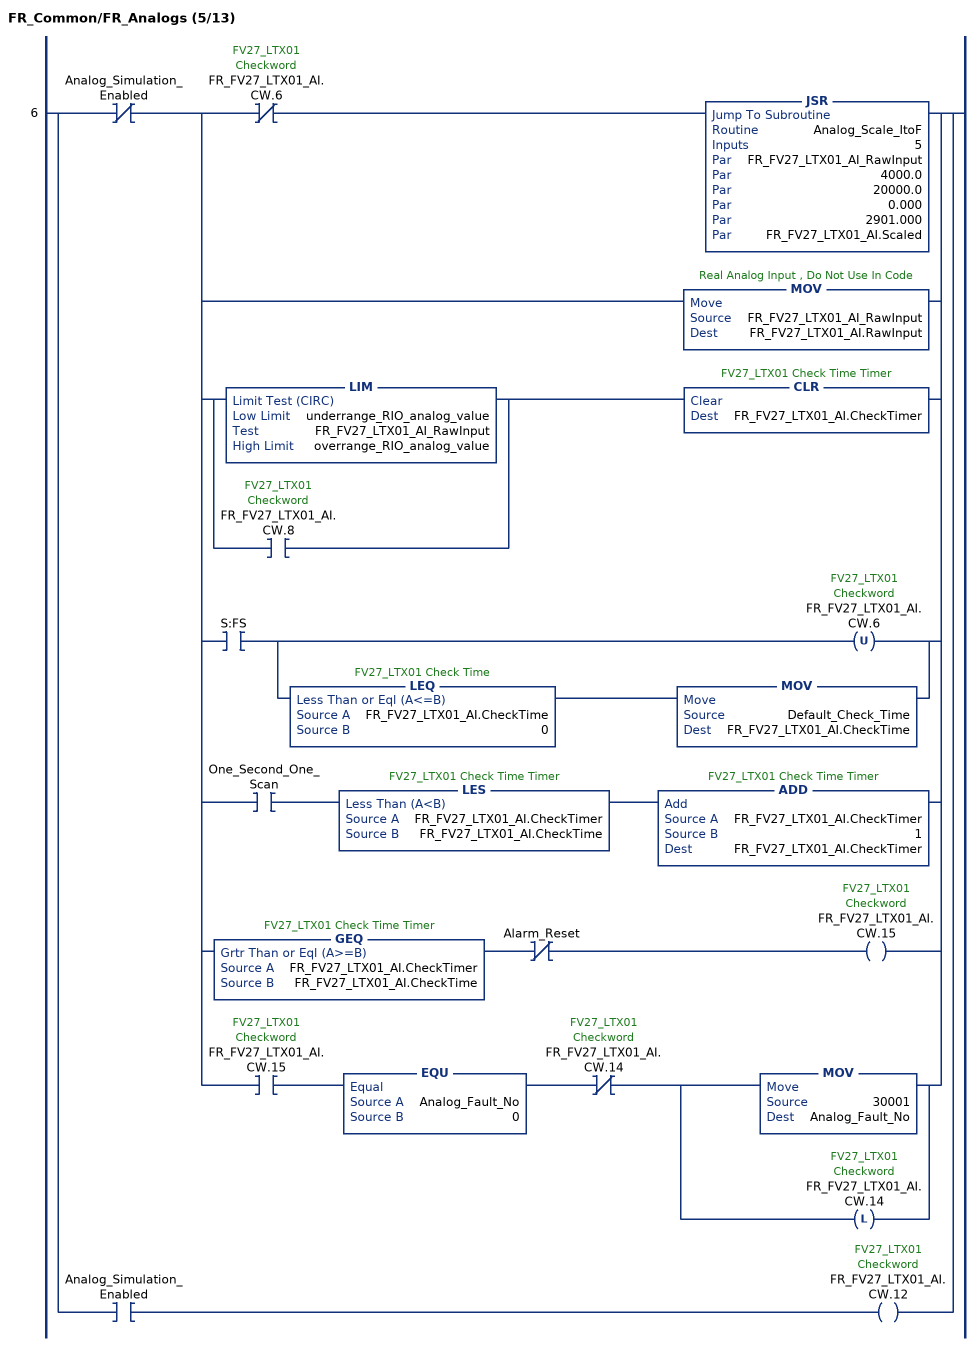
   6: [XIO(Analog_Simulation_Enabled) [XIO(FR_FV27_LTX01_AI.CW.6) JSR(Analog_Scale_ItoF,5,FR_FV27_LTX01_AI_RawInput,4000.0,20000.0,0.000,2901.000,FR_FV27_LTX01_AI.Scaled) ,MOV(FR_FV27_LTX01_AI_RawInput,FR_FV27_LTX01_AI.RawInput) ,[LIM(underrange_RIO_analog_value,FR_FV27_LTX01_AI_RawInput,overrange_RIO_analog_value) ,XIC(FR_FV27_LTX01_AI.CW.8) ] CLR(FR_FV27_LTX01_AI.CheckTimer) ,XIC(S:FS) [OTU(FR_FV27_LTX01_AI.CW.6) ,LEQ(FR_FV27_LTX01_AI.CheckTime,0) MOV(Default_Check_Time,FR_FV27_LTX01_AI.CheckTime) ] ,XIC(One_Second_One_Scan) LES(FR_FV27_LTX01_AI.CheckTimer,FR_FV27_LTX01_AI.CheckTime) ADD(FR_FV27_LTX01_AI.CheckTimer,1,FR_FV27_LTX01_AI.CheckTimer) ,GEQ(FR_FV27_LTX01_AI.CheckTimer,FR_FV27_LTX01_AI.CheckTime) XIO(Alarm_Reset) OTE(FR_FV27_LTX01_AI.CW.15) ,XIC(FR_FV27_LTX01_AI.CW.15) EQU(Analog_Fault_No,0) XIO(FR_FV27_LTX01_AI.CW.14) [MOV(30001,Analog_Fault_No) ,OTL(FR_FV27_LTX01_AI.CW.14) ] ] ,XIC(Analog_Simulation_Enabled) OTE(FR_FV27_LTX01_AI.CW.12) ];
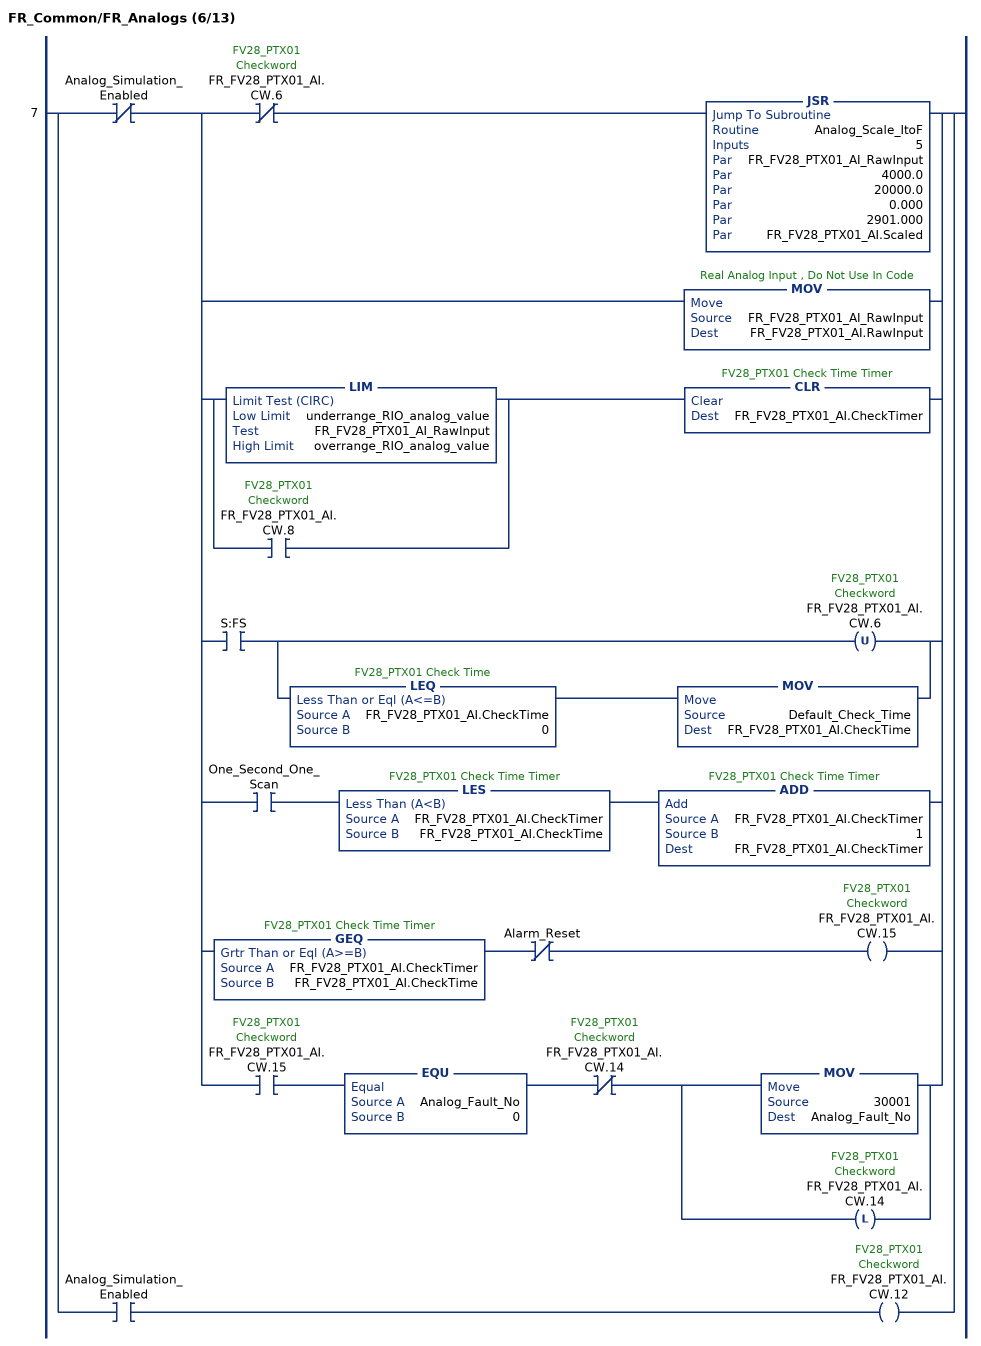
   7: [XIO(Analog_Simulation_Enabled) [XIO(FR_FV28_PTX01_AI.CW.6) JSR(Analog_Scale_ItoF,5,FR_FV28_PTX01_AI_RawInput,4000.0,20000.0,0.000,2901.000,FR_FV28_PTX01_AI.Scaled) ,MOV(FR_FV28_PTX01_AI_RawInput,FR_FV28_PTX01_AI.RawInput) ,[LIM(underrange_RIO_analog_value,FR_FV28_PTX01_AI_RawInput,overrange_RIO_analog_value) ,XIC(FR_FV28_PTX01_AI.CW.8) ] CLR(FR_FV28_PTX01_AI.CheckTimer) ,XIC(S:FS) [OTU(FR_FV28_PTX01_AI.CW.6) ,LEQ(FR_FV28_PTX01_AI.CheckTime,0) MOV(Default_Check_Time,FR_FV28_PTX01_AI.CheckTime) ] ,XIC(One_Second_One_Scan) LES(FR_FV28_PTX01_AI.CheckTimer,FR_FV28_PTX01_AI.CheckTime) ADD(FR_FV28_PTX01_AI.CheckTimer,1,FR_FV28_PTX01_AI.CheckTimer) ,GEQ(FR_FV28_PTX01_AI.CheckTimer,FR_FV28_PTX01_AI.CheckTime) XIO(Alarm_Reset) OTE(FR_FV28_PTX01_AI.CW.15) ,XIC(FR_FV28_PTX01_AI.CW.15) EQU(Analog_Fault_No,0) XIO(FR_FV28_PTX01_AI.CW.14) [MOV(30001,Analog_Fault_No) ,OTL(FR_FV28_PTX01_AI.CW.14) ] ] ,XIC(Analog_Simulation_Enabled) OTE(FR_FV28_PTX01_AI.CW.12) ];
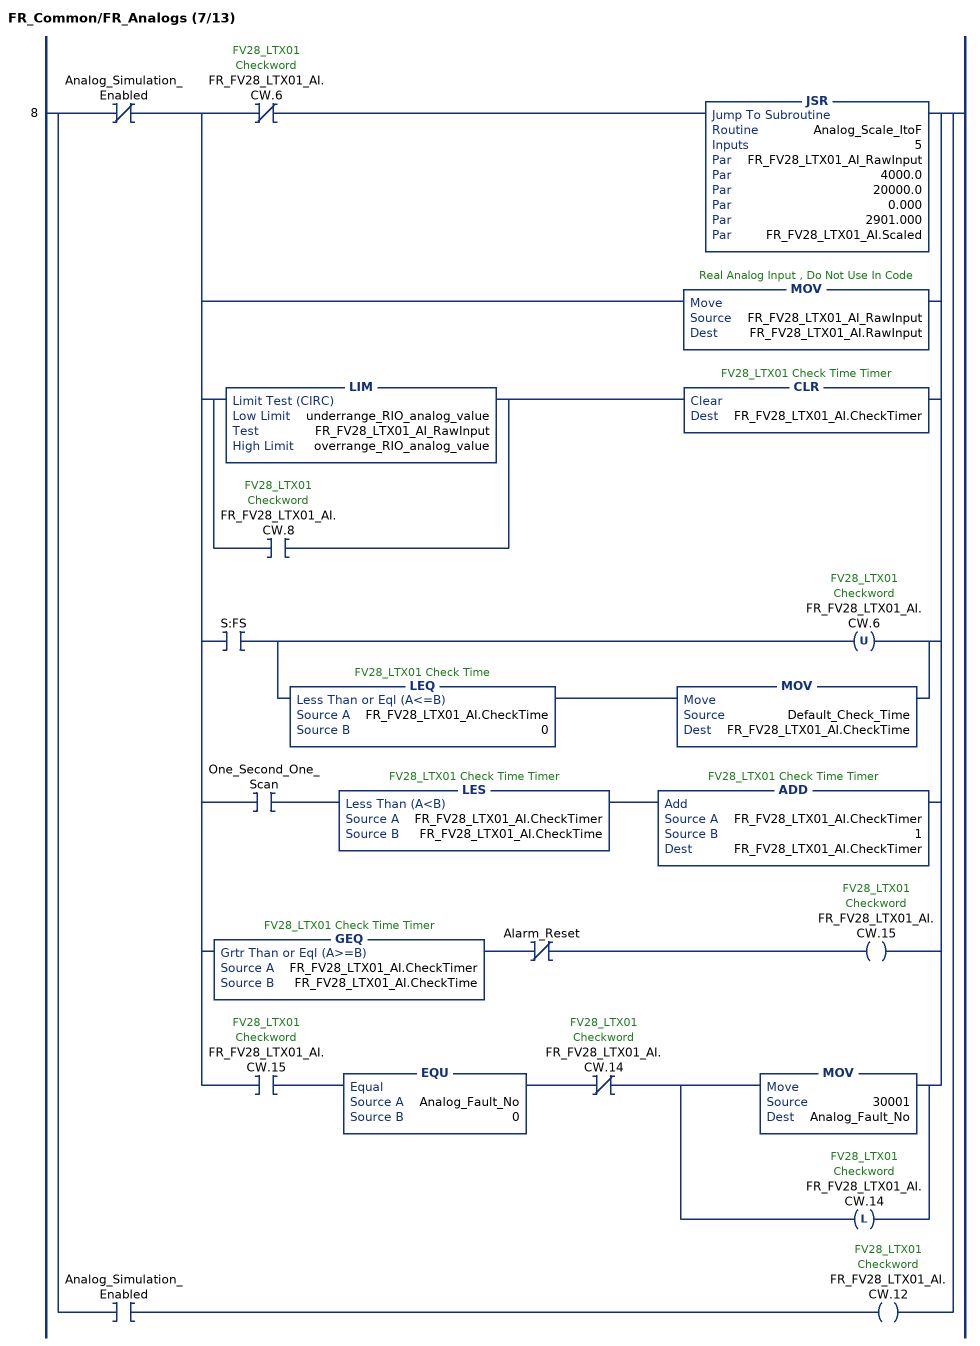
   8: [XIO(Analog_Simulation_Enabled) [XIO(FR_FV28_LTX01_AI.CW.6) JSR(Analog_Scale_ItoF,5,FR_FV28_LTX01_AI_RawInput,4000.0,20000.0,0.000,2901.000,FR_FV28_LTX01_AI.Scaled) ,MOV(FR_FV28_LTX01_AI_RawInput,FR_FV28_LTX01_AI.RawInput) ,[LIM(underrange_RIO_analog_value,FR_FV28_LTX01_AI_RawInput,overrange_RIO_analog_value) ,XIC(FR_FV28_LTX01_AI.CW.8) ] CLR(FR_FV28_LTX01_AI.CheckTimer) ,XIC(S:FS) [OTU(FR_FV28_LTX01_AI.CW.6) ,LEQ(FR_FV28_LTX01_AI.CheckTime,0) MOV(Default_Check_Time,FR_FV28_LTX01_AI.CheckTime) ] ,XIC(One_Second_One_Scan) LES(FR_FV28_LTX01_AI.CheckTimer,FR_FV28_LTX01_AI.CheckTime) ADD(FR_FV28_LTX01_AI.CheckTimer,1,FR_FV28_LTX01_AI.CheckTimer) ,GEQ(FR_FV28_LTX01_AI.CheckTimer,FR_FV28_LTX01_AI.CheckTime) XIO(Alarm_Reset) OTE(FR_FV28_LTX01_AI.CW.15) ,XIC(FR_FV28_LTX01_AI.CW.15) EQU(Analog_Fault_No,0) XIO(FR_FV28_LTX01_AI.CW.14) [MOV(30001,Analog_Fault_No) ,OTL(FR_FV28_LTX01_AI.CW.14) ] ] ,XIC(Analog_Simulation_Enabled) OTE(FR_FV28_LTX01_AI.CW.12) ];
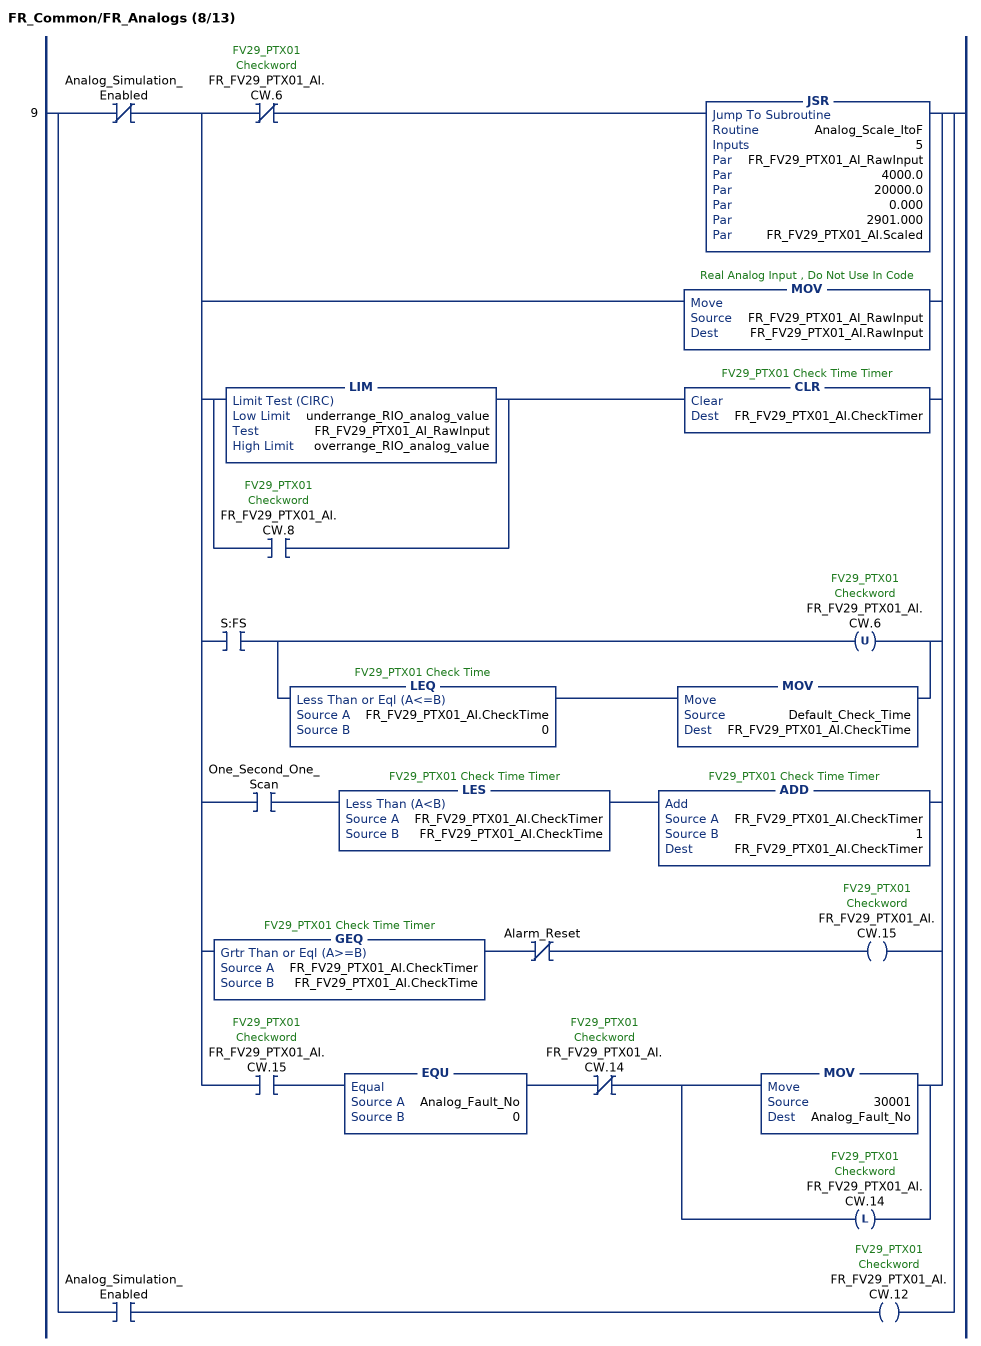
   9: [XIO(Analog_Simulation_Enabled) [XIO(FR_FV29_PTX01_AI.CW.6) JSR(Analog_Scale_ItoF,5,FR_FV29_PTX01_AI_RawInput,4000.0,20000.0,0.000,2901.000,FR_FV29_PTX01_AI.Scaled) ,MOV(FR_FV29_PTX01_AI_RawInput,FR_FV29_PTX01_AI.RawInput) ,[LIM(underrange_RIO_analog_value,FR_FV29_PTX01_AI_RawInput,overrange_RIO_analog_value) ,XIC(FR_FV29_PTX01_AI.CW.8) ] CLR(FR_FV29_PTX01_AI.CheckTimer) ,XIC(S:FS) [OTU(FR_FV29_PTX01_AI.CW.6) ,LEQ(FR_FV29_PTX01_AI.CheckTime,0) MOV(Default_Check_Time,FR_FV29_PTX01_AI.CheckTime) ] ,XIC(One_Second_One_Scan) LES(FR_FV29_PTX01_AI.CheckTimer,FR_FV29_PTX01_AI.CheckTime) ADD(FR_FV29_PTX01_AI.CheckTimer,1,FR_FV29_PTX01_AI.CheckTimer) ,GEQ(FR_FV29_PTX01_AI.CheckTimer,FR_FV29_PTX01_AI.CheckTime) XIO(Alarm_Reset) OTE(FR_FV29_PTX01_AI.CW.15) ,XIC(FR_FV29_PTX01_AI.CW.15) EQU(Analog_Fault_No,0) XIO(FR_FV29_PTX01_AI.CW.14) [MOV(30001,Analog_Fault_No) ,OTL(FR_FV29_PTX01_AI.CW.14) ] ] ,XIC(Analog_Simulation_Enabled) OTE(FR_FV29_PTX01_AI.CW.12) ];
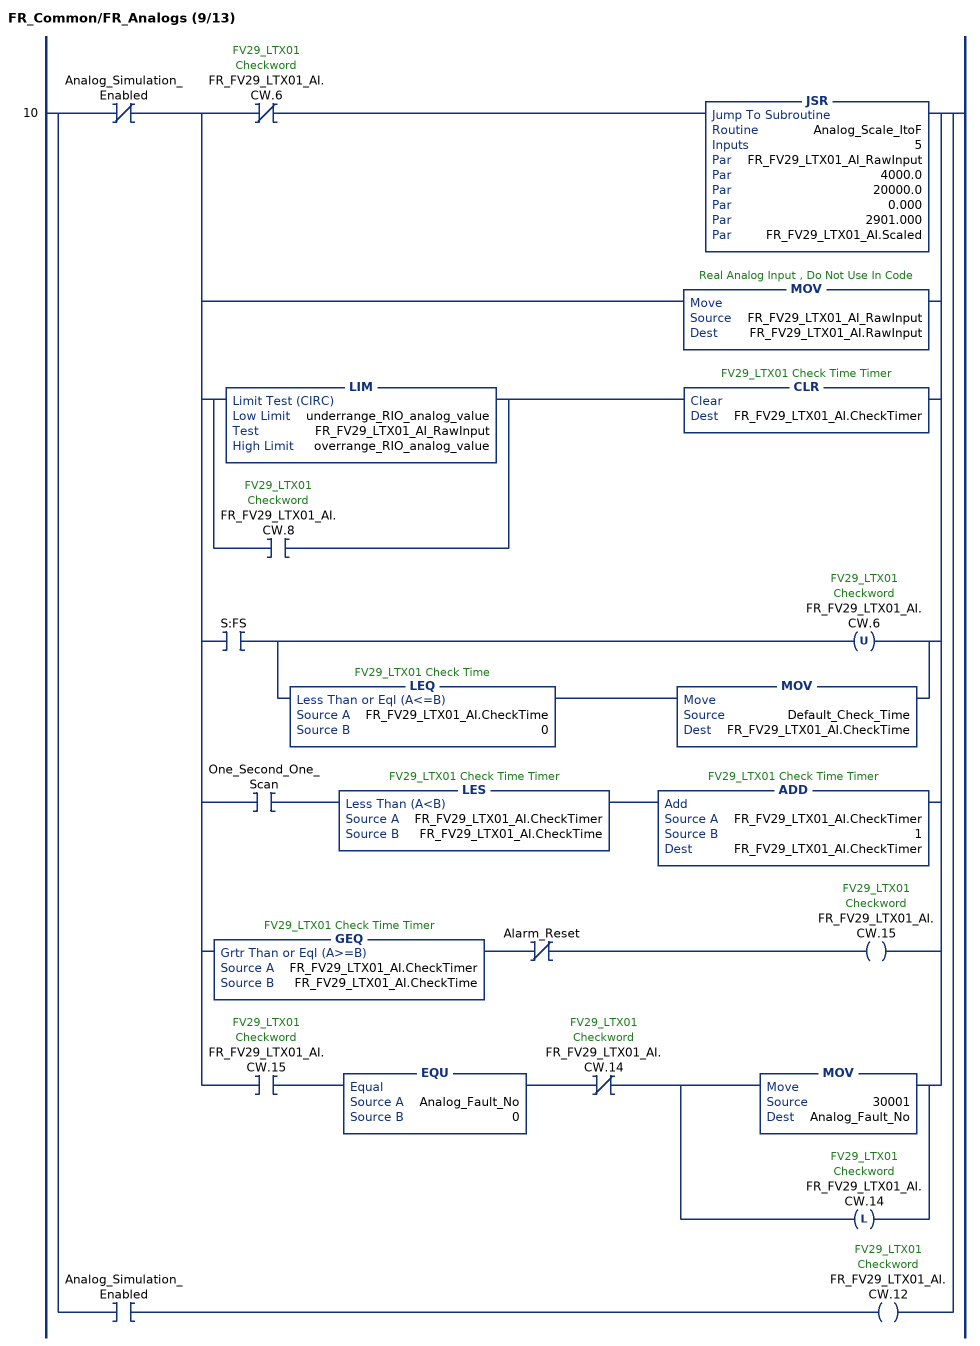
   10: [XIO(Analog_Simulation_Enabled) [XIO(FR_FV29_LTX01_AI.CW.6) JSR(Analog_Scale_ItoF,5,FR_FV29_LTX01_AI_RawInput,4000.0,20000.0,0.000,2901.000,FR_FV29_LTX01_AI.Scaled) ,MOV(FR_FV29_LTX01_AI_RawInput,FR_FV29_LTX01_AI.RawInput) ,[LIM(underrange_RIO_analog_value,FR_FV29_LTX01_AI_RawInput,overrange_RIO_analog_value) ,XIC(FR_FV29_LTX01_AI.CW.8) ] CLR(FR_FV29_LTX01_AI.CheckTimer) ,XIC(S:FS) [OTU(FR_FV29_LTX01_AI.CW.6) ,LEQ(FR_FV29_LTX01_AI.CheckTime,0) MOV(Default_Check_Time,FR_FV29_LTX01_AI.CheckTime) ] ,XIC(One_Second_One_Scan) LES(FR_FV29_LTX01_AI.CheckTimer,FR_FV29_LTX01_AI.CheckTime) ADD(FR_FV29_LTX01_AI.CheckTimer,1,FR_FV29_LTX01_AI.CheckTimer) ,GEQ(FR_FV29_LTX01_AI.CheckTimer,FR_FV29_LTX01_AI.CheckTime) XIO(Alarm_Reset) OTE(FR_FV29_LTX01_AI.CW.15) ,XIC(FR_FV29_LTX01_AI.CW.15) EQU(Analog_Fault_No,0) XIO(FR_FV29_LTX01_AI.CW.14) [MOV(30001,Analog_Fault_No) ,OTL(FR_FV29_LTX01_AI.CW.14) ] ] ,XIC(Analog_Simulation_Enabled) OTE(FR_FV29_LTX01_AI.CW.12) ];
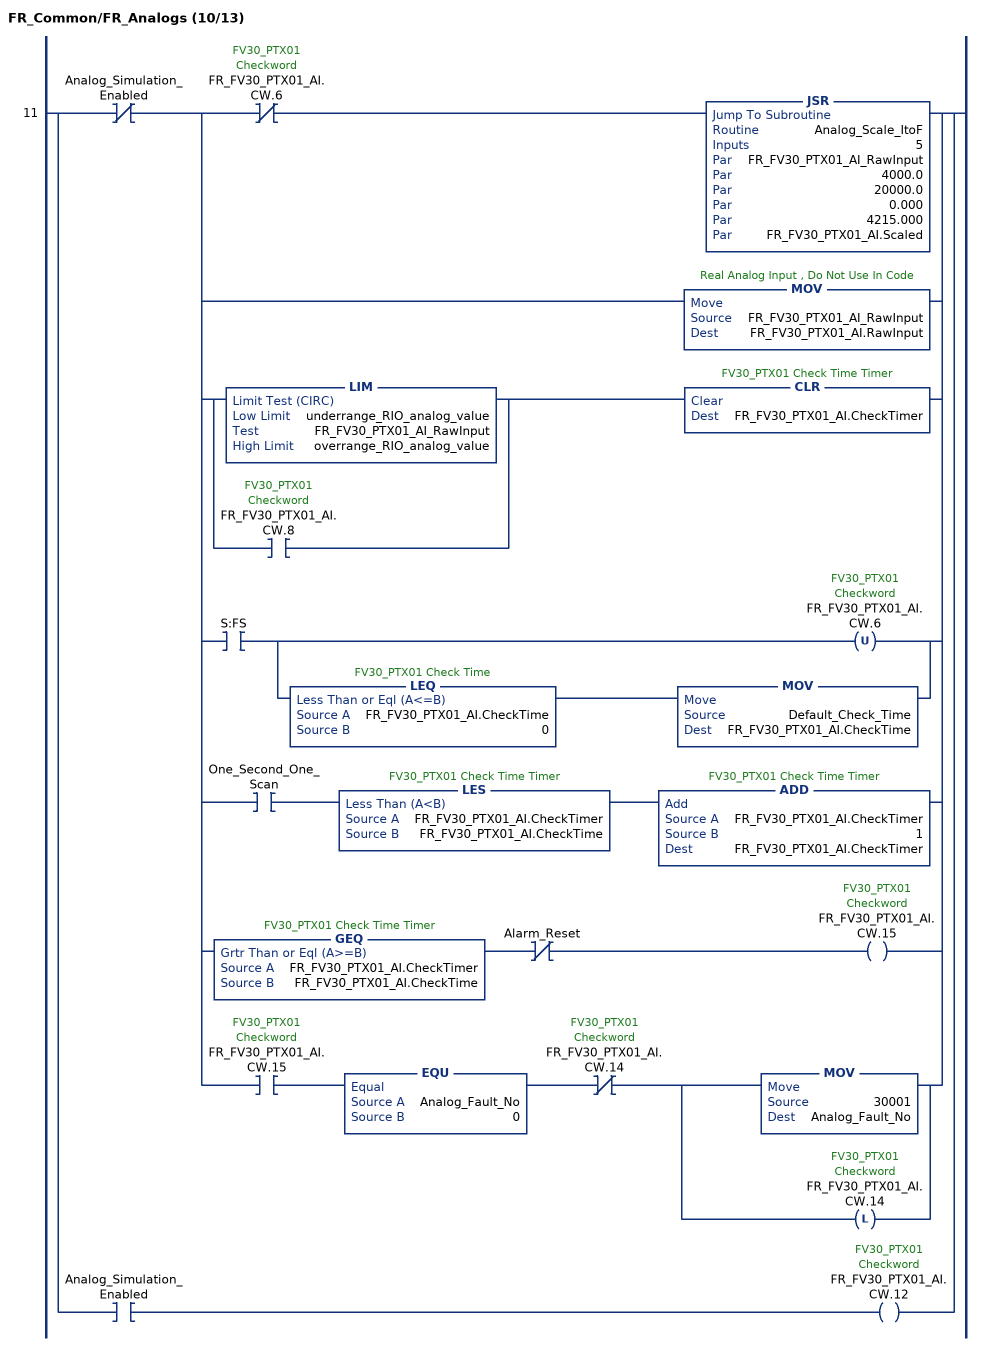
   11: [XIO(Analog_Simulation_Enabled) [XIO(FR_FV30_PTX01_AI.CW.6) JSR(Analog_Scale_ItoF,5,FR_FV30_PTX01_AI_RawInput,4000.0,20000.0,0.000,4215.000,FR_FV30_PTX01_AI.Scaled) ,MOV(FR_FV30_PTX01_AI_RawInput,FR_FV30_PTX01_AI.RawInput) ,[LIM(underrange_RIO_analog_value,FR_FV30_PTX01_AI_RawInput,overrange_RIO_analog_value) ,XIC(FR_FV30_PTX01_AI.CW.8) ] CLR(FR_FV30_PTX01_AI.CheckTimer) ,XIC(S:FS) [OTU(FR_FV30_PTX01_AI.CW.6) ,LEQ(FR_FV30_PTX01_AI.CheckTime,0) MOV(Default_Check_Time,FR_FV30_PTX01_AI.CheckTime) ] ,XIC(One_Second_One_Scan) LES(FR_FV30_PTX01_AI.CheckTimer,FR_FV30_PTX01_AI.CheckTime) ADD(FR_FV30_PTX01_AI.CheckTimer,1,FR_FV30_PTX01_AI.CheckTimer) ,GEQ(FR_FV30_PTX01_AI.CheckTimer,FR_FV30_PTX01_AI.CheckTime) XIO(Alarm_Reset) OTE(FR_FV30_PTX01_AI.CW.15) ,XIC(FR_FV30_PTX01_AI.CW.15) EQU(Analog_Fault_No,0) XIO(FR_FV30_PTX01_AI.CW.14) [MOV(30001,Analog_Fault_No) ,OTL(FR_FV30_PTX01_AI.CW.14) ] ] ,XIC(Analog_Simulation_Enabled) OTE(FR_FV30_PTX01_AI.CW.12) ];
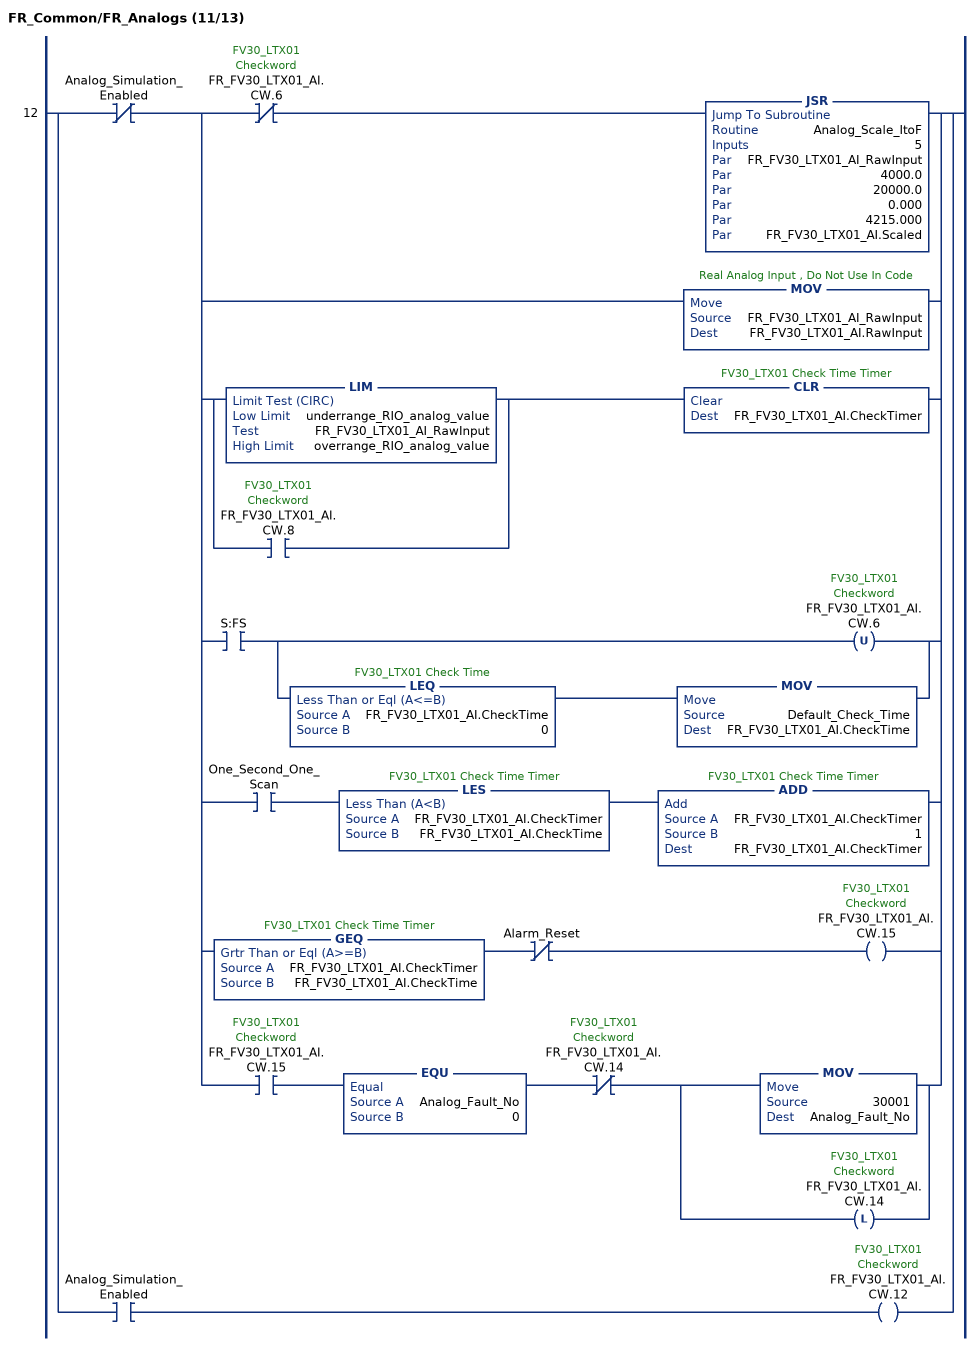
   12: [XIO(Analog_Simulation_Enabled) [XIO(FR_FV30_LTX01_AI.CW.6) JSR(Analog_Scale_ItoF,5,FR_FV30_LTX01_AI_RawInput,4000.0,20000.0,0.000,4215.000,FR_FV30_LTX01_AI.Scaled) ,MOV(FR_FV30_LTX01_AI_RawInput,FR_FV30_LTX01_AI.RawInput) ,[LIM(underrange_RIO_analog_value,FR_FV30_LTX01_AI_RawInput,overrange_RIO_analog_value) ,XIC(FR_FV30_LTX01_AI.CW.8) ] CLR(FR_FV30_LTX01_AI.CheckTimer) ,XIC(S:FS) [OTU(FR_FV30_LTX01_AI.CW.6) ,LEQ(FR_FV30_LTX01_AI.CheckTime,0) MOV(Default_Check_Time,FR_FV30_LTX01_AI.CheckTime) ] ,XIC(One_Second_One_Scan) LES(FR_FV30_LTX01_AI.CheckTimer,FR_FV30_LTX01_AI.CheckTime) ADD(FR_FV30_LTX01_AI.CheckTimer,1,FR_FV30_LTX01_AI.CheckTimer) ,GEQ(FR_FV30_LTX01_AI.CheckTimer,FR_FV30_LTX01_AI.CheckTime) XIO(Alarm_Reset) OTE(FR_FV30_LTX01_AI.CW.15) ,XIC(FR_FV30_LTX01_AI.CW.15) EQU(Analog_Fault_No,0) XIO(FR_FV30_LTX01_AI.CW.14) [MOV(30001,Analog_Fault_No) ,OTL(FR_FV30_LTX01_AI.CW.14) ] ] ,XIC(Analog_Simulation_Enabled) OTE(FR_FV30_LTX01_AI.CW.12) ];
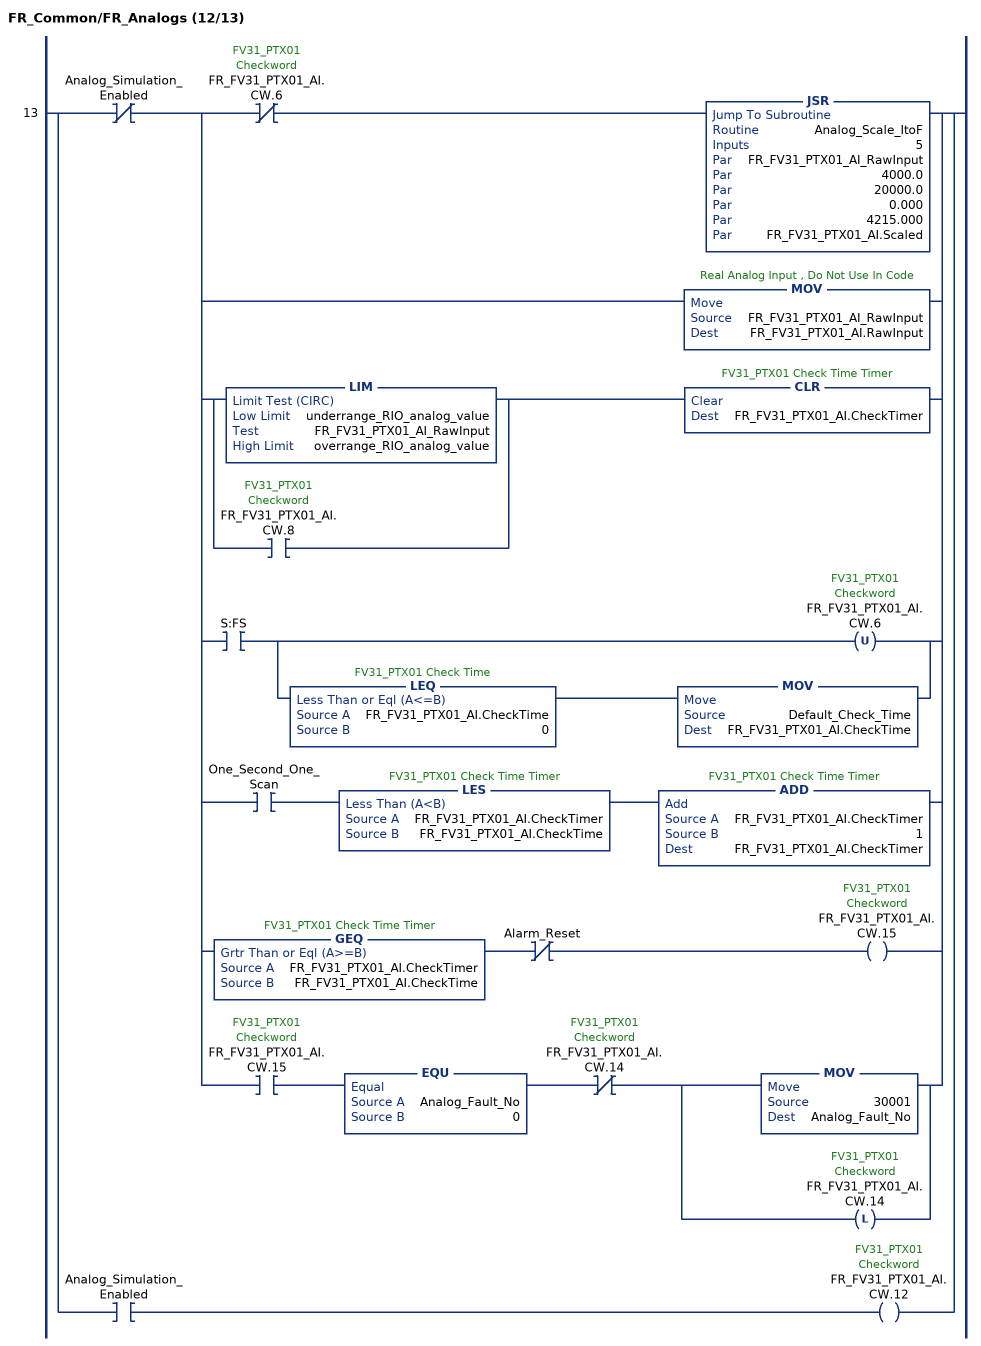
   13: [XIO(Analog_Simulation_Enabled) [XIO(FR_FV31_PTX01_AI.CW.6) JSR(Analog_Scale_ItoF,5,FR_FV31_PTX01_AI_RawInput,4000.0,20000.0,0.000,4215.000,FR_FV31_PTX01_AI.Scaled) ,MOV(FR_FV31_PTX01_AI_RawInput,FR_FV31_PTX01_AI.RawInput) ,[LIM(underrange_RIO_analog_value,FR_FV31_PTX01_AI_RawInput,overrange_RIO_analog_value) ,XIC(FR_FV31_PTX01_AI.CW.8) ] CLR(FR_FV31_PTX01_AI.CheckTimer) ,XIC(S:FS) [OTU(FR_FV31_PTX01_AI.CW.6) ,LEQ(FR_FV31_PTX01_AI.CheckTime,0) MOV(Default_Check_Time,FR_FV31_PTX01_AI.CheckTime) ] ,XIC(One_Second_One_Scan) LES(FR_FV31_PTX01_AI.CheckTimer,FR_FV31_PTX01_AI.CheckTime) ADD(FR_FV31_PTX01_AI.CheckTimer,1,FR_FV31_PTX01_AI.CheckTimer) ,GEQ(FR_FV31_PTX01_AI.CheckTimer,FR_FV31_PTX01_AI.CheckTime) XIO(Alarm_Reset) OTE(FR_FV31_PTX01_AI.CW.15) ,XIC(FR_FV31_PTX01_AI.CW.15) EQU(Analog_Fault_No,0) XIO(FR_FV31_PTX01_AI.CW.14) [MOV(30001,Analog_Fault_No) ,OTL(FR_FV31_PTX01_AI.CW.14) ] ] ,XIC(Analog_Simulation_Enabled) OTE(FR_FV31_PTX01_AI.CW.12) ];
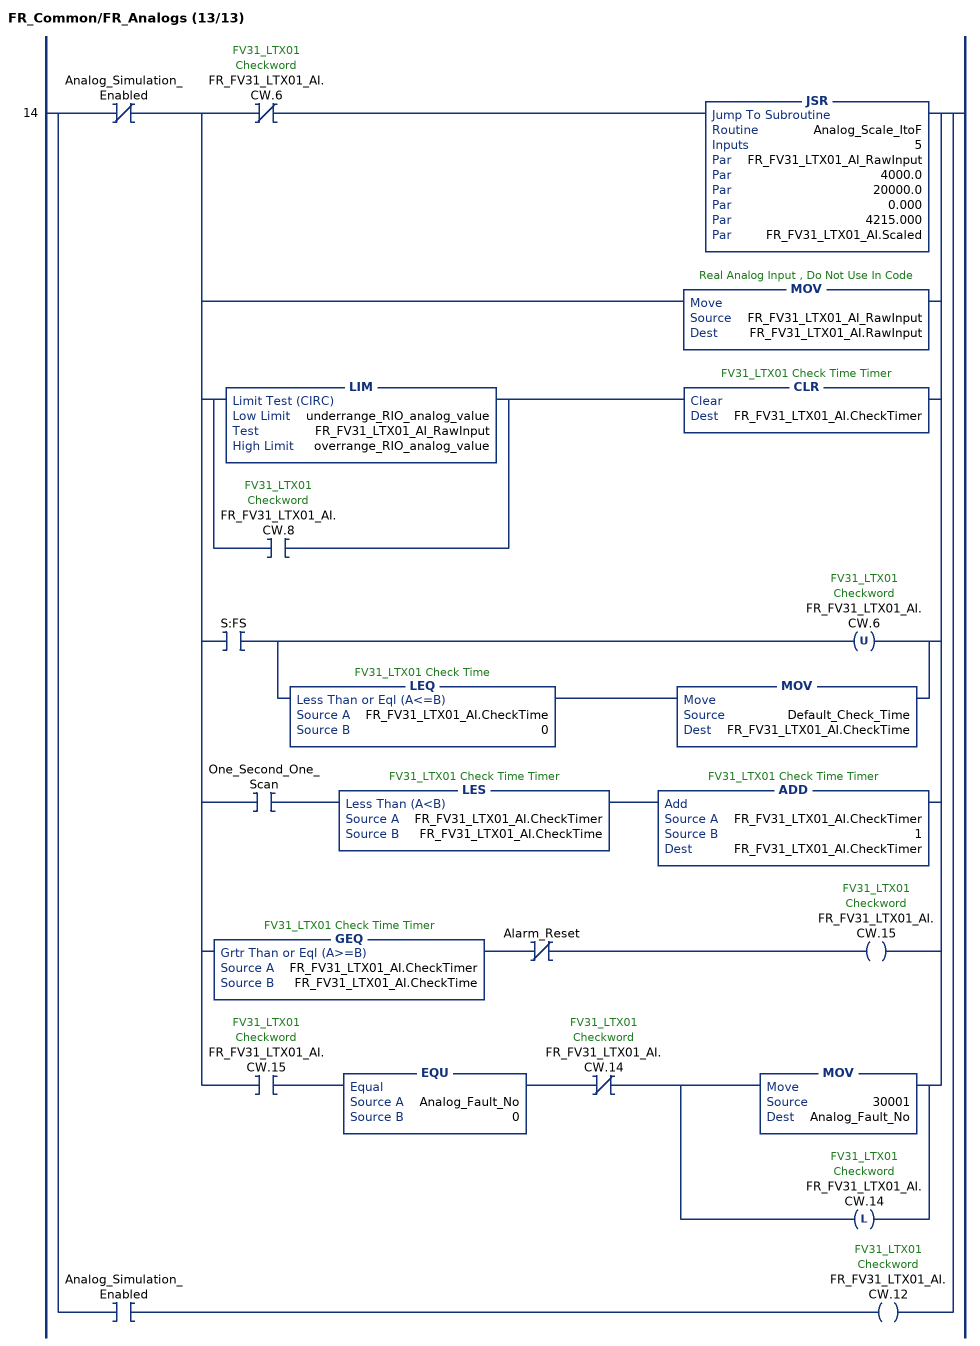
   14: [XIO(Analog_Simulation_Enabled) [XIO(FR_FV31_LTX01_AI.CW.6) JSR(Analog_Scale_ItoF,5,FR_FV31_LTX01_AI_RawInput,4000.0,20000.0,0.000,4215.000,FR_FV31_LTX01_AI.Scaled) ,MOV(FR_FV31_LTX01_AI_RawInput,FR_FV31_LTX01_AI.RawInput) ,[LIM(underrange_RIO_analog_value,FR_FV31_LTX01_AI_RawInput,overrange_RIO_analog_value) ,XIC(FR_FV31_LTX01_AI.CW.8) ] CLR(FR_FV31_LTX01_AI.CheckTimer) ,XIC(S:FS) [OTU(FR_FV31_LTX01_AI.CW.6) ,LEQ(FR_FV31_LTX01_AI.CheckTime,0) MOV(Default_Check_Time,FR_FV31_LTX01_AI.CheckTime) ] ,XIC(One_Second_One_Scan) LES(FR_FV31_LTX01_AI.CheckTimer,FR_FV31_LTX01_AI.CheckTime) ADD(FR_FV31_LTX01_AI.CheckTimer,1,FR_FV31_LTX01_AI.CheckTimer) ,GEQ(FR_FV31_LTX01_AI.CheckTimer,FR_FV31_LTX01_AI.CheckTime) XIO(Alarm_Reset) OTE(FR_FV31_LTX01_AI.CW.15) ,XIC(FR_FV31_LTX01_AI.CW.15) EQU(Analog_Fault_No,0) XIO(FR_FV31_LTX01_AI.CW.14) [MOV(30001,Analog_Fault_No) ,OTL(FR_FV31_LTX01_AI.CW.14) ] ] ,XIC(Analog_Simulation_Enabled) OTE(FR_FV31_LTX01_AI.CW.12) ];
END_ROUTINE
